// Mitsubishi GX Works2 project: ZhaoQing_HuaCheng1_Debug   PLC: Q06UDEH (continued)
    
    IF Import2Conveyor2IO.xEmpty=0 AND XF5 THEN
    	Import2LoadCylinderIO.xMDIExe:=1;
    	Import2LoadCylinderIO.iDestinationPos:=2;
    	Import2Conveyor2IO.xPutInto:=0;
    END_IF;
    IF NOT XF5 THEN
    	Import2LoadCylinderIO.xMDIExe:=1;
    	Import2LoadCylinderIO.iDestinationPos:=1;	
    END_IF;
    IF LDP(TRUE, Import2LoadCylinderIO.iCurrentPos=1) THEN
    	Import2Conveyor2IO.xPutInto:=1;
    END_IF;
   (*空框回流*)
    (*A内衬空框回流*) 
   IF  LDP(TRUE,H2200Switch1TaskID=1) THEN
   	m_xCartonADischargeLock:=1;(*A内衬空框回流下料锁，保证一次下料任务只下一个料*) 
   END_IF;
   IF LDF(TRUE,H2200BayCylinderEmptyABackIO.xUnload) OR H2200Switch1TaskID=0  THEN
   	m_xCartonADischargeLock:=0;
   END_IF;
   H2200BayCylinderEmptyABackIO.xUnload:=H2200SwitchEmptyABackConveyorIn.xEmpty
   																				 AND  H2200Switch1ConveyorIn.xEmpty
   																				 AND m_xCartonADischargeLock;
   H2200SwitchEmptyABackIO.xEntryEnable:=H2200BayCylinderEmptyABackIO.xNextRun;
   H2200SwitchEmptyABackIO.xLiftCylinderExtendInit:=H2200Switch1TaskID=1;
    H2200SwitchEmptyABackIO.xSwithEnable:=1;
    (*B内衬空框回流*) 
    IF  LDP(TRUE,H2200Switch1TaskID=2) THEN
   	m_xCartonBDischargeLock:=1;(*B内衬空框回流下料锁，保证一次下料任务只下一个料*) 
   END_IF;
   IF LDF(TRUE,H2200BayCylinderEmptyBBackIO.xUnload) OR H2200Switch1TaskID=0  THEN
   	m_xCartonBDischargeLock:=0;
   END_IF;
   H2200BayCylinderEmptyBBackIO.xUnload:=H2200SwitchEmptyBBackConveyorIn.xEmpty 
   																				 AND  H2200Switch1ConveyorIn.xEmpty
   																				 AND m_xCartonBDischargeLock;
   H2200SwitchEmptyBBackIO.xEntryEnable:=H2200BayCylinderEmptyBBackIO.xNextRun;
   H2200SwitchEmptyBBackIO.xLiftCylinderExtendInit:=1;
    H2200SwitchEmptyBBackIO.xSwithEnable:=1;    
    (*H2200Switch1 空框去注液任务*)
    IF H2200Switch1TaskID=1 OR H2200Switch1TaskID=2  THEN
    	H2200SwitchEmptyABackIO.xExitEnable:=H2200Switch1ConveyorIn.xEmpty; 
    	H2200SwitchEmptyBBackIO.xExitEnable:=H2200Switch1ConveyorIn.xEmpty;   	
    	H2200Switch1IO.xEntryEnable:=H2200SwitchEmptyABackConveyorOut.xNextRun OR H2200SwitchEmptyBBackConveyorOut.xNextRun ;
    	H2200Switch1IO.xSwithEnable:=0;
    	H2200Switch1IO.xExitEnable:=H2200RotorConveyorIO.xEmpty AND H2200RotorIO.iCurrentPos=1 AND X75;
    ELSE
    	H2200Switch1IO.xEntryEnable:=0;
    	H2200SwitchEmptyABackIO.xExitEnable:=0;
    	H2200SwitchEmptyBBackIO.xExitEnable:=0;
    	H2200Switch1IO.xExitEnable:=0;
    END_IF;
    (*H2200Switch1 满框入库任务*)
    IF H2200Switch1TaskID<>5 THEN
    	H2200Switch1IO.xLiftCylinderExtendInit:=0;
    END_IF;
    IF H2200RotorConveyorIO.xEmpty THEN
    	H2200RotorIO.xMDIExe:=1;
    	H2200RotorIO.iDestinationPos:=1;
    END_IF;
    IF H2200RotorConveyorIO.xEmpty=0 THEN
     	H2200RotorIO.xMDIExe:=1;
    	H2200RotorIO.iDestinationPos:=2;   
    END_IF;   
    IF H2200RotorIO.iCurrentPos=1 AND X75 THEN
    	H2200RotorConveyorIO.xLoad:=H2200Switch1ConveyorIn.xNextRun;
    ELSE
    	H2200RotorConveyorIO.xLoad:=0;	
    END_IF;
    IF Conveyor1IO.xEmpty THEN
    	Lifter1IO.xMDIExe:=1;
    	Lifter1IO.iDestinationPos:=2;
    END_IF;
    IF Conveyor1IO.xEmpty=0 THEN
    	Lifter1IO.xMDIExe:=1;
    	Lifter1IO.iDestinationPos:=1; 
    END_IF;
    H2200RotorConveyorIO.xUnloadCCW:=1;
    IF Lifter1IO.iCurrentPos=2 AND X8D AND H2200RotorIO.iCurrentPos=2 AND X6F THEN
    	H2200RotorConveyorIO.xUnload:=Conveyor1IO.xEmpty;
    ELSE
    	H2200RotorConveyorIO.xUnload:=0;
    END_IF;
    Conveyor1IO.xLoad:=H2200RotorConveyorIO.xNextRun; 
    IF Lifter1IO.iCurrentPos=1 AND X8C THEN
    	Conveyor1IO.xUnload:=H850Conveyor3IO.xEmpty;
    ELSE
    	Conveyor1IO.xUnload:=0;
    END_IF;  	
    H850Conveyor3IO.xLoad:=Conveyor1IO.xNextRun;
    h850conveyor3IO.xUnload:=H850Conveyor1IO.xEmpty;
    H850Conveyor1IO.xLoad:=H850Conveyor3IO.xNextRun;
    H850Conveyor1IO.xPutInto:=NOT H850Conveyor1IO.xBusy AND  SM412;
END_IF;
Y1B1:=M134 AND g_xEStop;(*空框A回流倍速链*)
Y1B0:=M135 AND g_xEStop;(*空框B回流倍速链*)
IF g_xManual THEN
    D201:=0;(*发送给化成B柜*)
    (************发送给上位机程序复位**************)
    D3100:=0;
    D3105:=0;
    D3120:=0;
    D3125:=0;
    D3016:=0;
    D3011:=0;
    D3300:=0;
    D3305:=0;
    D3310:=0;
    (*****************************************************)
	IF M163 THEN (*入库倍速链 手动*)
		 Y186:=1;(*入库倍速链*)
	ELSE
		Y186:=0;(*入库倍速链*)
	END_IF;
	IF M64 THEN (*出库倍速链 手动*)
		 Y187:=1;(*出库倍速链 *)
	ELSE
		Y187:=0;(*出库倍速链 *)
	END_IF;		
END_IF;


    (*报警*)
    M300:=NOT H3000SwitchPackageConveyorIn.xEmpty;
    M301:=H3000SwitchPackageConveyorIn.xUnloadAlarm;
    M302:=NOT H3000SwitchPackageConveyorOut.xEmpty;
    M303:=H3000SwitchPackageConveyorOut.xUnloadAlarm;   
    M304:=NOT H3000SwitchChemConveyorIn.xEmpty;
    M305:=H3000SwitchChemConveyorIn.xUnloadAlarm;   
    M306:=NOT H3000SwitchChemConveyorOut.xEmpty;
    M307:=H3000SwitchChemConveyorOut.xUnloadAlarm;  
    M308:=NOT H3000Conveyor1IO.xEmpty;
    M309:=H3000Conveyor1IO.xUnloadAlarm;       
     M310:=NOT H3000Conveyor2IO.xEmpty;
    M311:=H3000Conveyor2IO.xUnloadAlarm;    
    M312:=NOT H3000Conveyor3IO.xEmpty;
    M313:=H3000Conveyor3IO.xUnloadAlarm; 
    M314:=NOT H3000Conveyor4IO.xEmpty;
    M315:=H3000Conveyor4IO.xUnloadAlarm;  
    M317:=NOT H3000Conveyor5IO.xEmpty;
    M318:=H3000Conveyor5IO.xUnloadAlarm; 
    M319:=NOT H3000Conveyor6IO.xEmpty;
    M320:=H3000Conveyor6IO.xUnloadAlarm;     
    M321:=NOT H3000Conveyor7IO.xEmpty;
    M322:=H3000Conveyor7IO.xUnloadAlarm;  
    M323:=NOT H3000Conveyor8IO.xEmpty;
    M324:=H3000Conveyor8IO.xUnloadAlarm;  
    M325:=NOT H3000Conveyor9IO.xEmpty;
    M326:=H3000Conveyor9IO.xUnloadAlarm;  
    M327:=NOT H3000Conveyor10IO.xEmpty;
    M328:=H3000Conveyor10IO.xUnloadAlarm;
    
    M329:=NOT H3000ChemConveyor2IO.xEmpty;
    M330:=H3000ChemConveyor2IO.xUnloadAlarm;
    M331:=NOT H3000ChemConveyor3IO.xEmpty;
    M332:=H3000ChemConveyor3IO.xUnloadAlarm;
    M333:=NOT H2200Switch1ConveyorIn.xEmpty;
    M334:=H2200Switch1ConveyorIn.xUnloadAlarm;
    M335:=NOT H2200Switch1ConveyorOut.xEmpty;
    M336:=H2200Switch1ConveyorOut.xUnloadAlarm;
    M337:=NOT H2200Switch2ConveyorIn.xEmpty;
    M338:=H2200Switch2ConveyorIn.xUnloadAlarm;
    M339:=NOT H2200Switch2ConveyorOut.xEmpty;
(*    M340:=H2200Switch2ConveyorOut.xUnloadAlarm;*)
     M341:=NOT H2200Conveyor1IO.xEmpty;
    M342:=H2200Conveyor1IO.xUnloadAlarm;       
     M343:=NOT H2200Conveyor2IO.xEmpty;
    M344:=H2200Conveyor2IO.xUnloadAlarm;    
    M345:=NOT H2200Conveyor3IO.xEmpty;
    M346:=H2200Conveyor3IO.xUnloadAlarm; 
    M347:=NOT H2200Conveyor4IO.xEmpty;
    M348:=H2200Conveyor4IO.xUnloadAlarm;  
    M349:=NOT H2200Conveyor5IO.xEmpty;
    M350:=H2200Conveyor5IO.xUnloadAlarm; 
    M351:=NOT H2200Conveyor6IO.xEmpty;
    M352:=H2200Conveyor6IO.xUnloadAlarm;     
    M353:=NOT H2200Conveyor7IO.xEmpty;
    M354:=H2200Conveyor7IO.xUnloadAlarm;  
    M355:=NOT H2200Conveyor8IO.xEmpty;
    M356:=H2200Conveyor8IO.xUnloadAlarm;  
    M357:=NOT H2200Conveyor9IO.xEmpty;
    M358:=H2200Conveyor9IO.xUnloadAlarm;  
    M359:=NOT H2200Conveyor10IO.xEmpty;
    M360:=H2200Conveyor10IO.xUnloadAlarm;
    M361:=NOT H2200ImportConveyor1IO.xEmpty;
    M362:=H2200ImportConveyor1IO.xUnloadAlarm;
     M363:=NOT H2200ImportConveyor2IO.xEmpty;
    M364:=H2200ImportConveyor2IO.xUnloadAlarm;   
     M365:=NOT H2200ImportConveyor3IO.xEmpty;
    M366:=H2200ImportConveyor3IO.xUnloadAlarm;    
    M367:=NOT H850Conveyor1IO.xEmpty;
    M368:=H850Conveyor1IO.xUnloadAlarm;      
     M369:=NOT H850Conveyor3IO.xEmpty;
    M370:=H850Conveyor3IO.xUnloadAlarm;  
    M371:=NOT H850Conveyor4IO.xEmpty;
    M372:=H850Conveyor4IO.xUnloadAlarm;
    M373:=NOT H850Conveyor5IO.xEmpty;
    M374:=H850Conveyor5IO.xUnloadAlarm;
    M375:=NOT H850Conveyor6IO.xEmpty;
    M376:=H850Conveyor6IO.xUnloadAlarm;
    M377:=NOT H850Conveyor7IO.xEmpty;
    M378:=H850Conveyor7IO.xUnloadAlarm; 
    M379:=NOT H850Conveyor8IO.xEmpty;
    M380:=H850Conveyor8IO.xUnloadAlarm; 
    M381:=NOT H850RotorConveyorIO.xEmpty;
    M382:=H850RotorConveyorIO.xUnloadAlarm;     
     
    M383:=D2335=1;(*化成入库后站台读码失败*)
    M384:=D2335=3;(*化成入库后站台条码重复*)
    M385:=D2340=1;(*注液入库前站台读码失败*)
    M386:=D2340=3;(*注液入库前站台条码重复*)
    M387:=D2300=1;(*高温入库分流读码失败*)
    M388:=D2305=1;(*高温出库分流读码失败*)
    M389:=D2310=1;(*提升机2分流读码失败*)
    M390:=Lifter2IO.xLooseAlarm;(*提升机2松绳检测*)
    M391:=Conveyor2IO.xOverWidthAlarm;(*提升机2超宽报警*)
    
    M392:=Import1SwitchConveyorOut.xUnloadAlarm;
    M393:=Import2SwitchConveyorOut.xUnloadAlarm;
    M394:=NOT H1000Conveyor1IO.xEmpty;
    M395:=H1000Conveyor1IO.xUnloadAlarm;
    M396:=NOT H1000Conveyor2IO.xEmpty;
    M397:=H1000Conveyor2IO.xUnloadAlarm;
    M398:=NOT H1000Conveyor3IO.xEmpty;
    M399:=H1000Conveyor3IO.xUnloadAlarm;
    M400:=NOT H1000Conveyor4IO.xEmpty;
    M401:=H1000Conveyor4IO.xUnloadAlarm;
    M402:=NOT H1000Conveyor5IO.xEmpty;
    M403:=H1000Conveyor5IO.xUnloadAlarm;
    M404:=NOT H1000Conveyor6IO.xEmpty;
    M405:=H1000Conveyor6IO.xUnloadAlarm;
    M406:=NOT H1000Conveyor7IO.xEmpty;
    M407:=H1000Conveyor7IO.xUnloadAlarm;
    M408:=NOT H1000Conveyor8IO.xEmpty;
    M409:=H1000Conveyor8IO.xUnloadAlarm;
    M410:=NOT H1000Conveyor9IO.xEmpty;
    M411:=H1000Conveyor9IO.xUnloadAlarm;
    M412:=NOT H1000Conveyor10IO.xEmpty;
    M413:=H1000Conveyor10IO.xUnloadAlarm;
    M414:=Export1Conveyor1IO.xUnloadAlarm;
    M415:= Export2Conveyor1IO.xUnloadAlarm;
     M416:=Export1Conveyor2IO.xUnloadAlarm;
    M417:= Export2Conveyor2IO.xUnloadAlarm;   
    M418:=H850SwitchConveyorOut.xUnloadAlarm;
    g_xAlarm:=M383 
    					OR M384 
    					OR M385 
    					OR M386 
    					OR M387 
    					OR M388 
    					OR M389 
    					OR M390 
    					OR M391 
    					OR  M307 
    					OR M382 
    					OR M392 
    					OR M393 
    					OR M362
    					OR M336
    					OR M414
    					OR M415
    					OR M416
    					OR M417
    					OR M418;
  IF LDP(TRUE, g_xManual) THEN
  	m_iExportConveyorOcuppy:=0;
  END_IF;
END_PROGRAM

FUNCTION_BLOCK PriorityFB
VAR_INPUT
  xCondition1 : BOOL;  (* 条件1 *)
  xCondition2 : BOOL;  (* 条件2 *)
  xCondition3 : BOOL;  (* 条件3 *)
  xCondition4 : BOOL;  (* 条件4 *)
  xCondition5 : BOOL;  (* 条件5 *)
  xTaskComplete : BOOL;  (* 任务完成 *)
  xReset : BOOL;  (* 复位 *)
END_VAR
VAR
  xOccupy : BOOL;  (* 占用 *)
END_VAR
VAR_OUTPUT
  iPriority : INT;  (* 输出任务号 *)
END_VAR
VAR
  m_tonConditionDelay : TON;
  m_xConditionDelay : BOOL;
  m_tConditionCurrentTime : TIME;
  m_iLastTask : INT;  (* 上次执行的任务 *)
  m_tpLastTaskPulse1 : TP;
  m_xLastTaskPulse : ARRAY [1..5] OF BOOL;
  m_tLastTaskPulse : ARRAY [1..5] OF TIME := [5(T#0s)];
  m_tpLastTaskPulse2 : TP;
  m_tpLastTaskPulse3 : TP;
  m_tpLastTaskPulse4 : TP;
  m_tpLastTaskPulse5 : TP;
END_VAR
(*我在reset那里加了Occupy的复位
任务为0时，Occupy也会自动复位
*)
IF NOT xCondition1 
	AND NOT xCondition2
	AND NOT xCondition3
	AND NOT xCondition4
	AND NOT xCondition5
	AND NOT xOccupy  THEN
	iPriority:=0;
END_IF;
IF LDP(TRUE, xTaskComplete) THEN
	xOccupy:=0;
	iPriority:=0;
END_IF;
m_tonConditionDelay(IN:= (xCondition1
                                                     OR  xCondition2
                                                     OR  xCondition3
                                                     OR  xCondition4
                                                     OR xCondition5)
                                                     AND iPriority=0,
                                                     PT:= T#1s,
                                                     Q:= m_xConditionDelay ,
                                                     ET:= m_tConditionCurrentTime );
m_tpLastTaskPulse1(IN:= xCondition1  AND m_iLastTask=1 AND m_xConditionDelay  ,PT:= T#1s,Q:= m_xLastTaskPulse[1],ET:= m_tLastTaskPulse[1] );
m_tpLastTaskPulse2(IN:= xCondition2  AND m_iLastTask=2 AND m_xConditionDelay,PT:= T#1s,Q:= m_xLastTaskPulse[2],ET:= m_tLastTaskPulse[2]);
m_tpLastTaskPulse3(IN:= xCondition3  AND m_iLastTask=3 AND m_xConditionDelay,PT:= T#1s,Q:= m_xLastTaskPulse[3],ET:= m_tLastTaskPulse[3] );
m_tpLastTaskPulse4(IN:= xCondition4  AND m_iLastTask=4 AND m_xConditionDelay,PT:= T#1s,Q:= m_xLastTaskPulse[4],ET:= m_tLastTaskPulse[4] );
m_tpLastTaskPulse5(IN:= xCondition5  AND m_iLastTask=5 AND m_xConditionDelay,PT:= T#1s,Q:= m_xLastTaskPulse[5],ET:= m_tLastTaskPulse[5] );

                                                     
IF xCondition1 AND NOT xOccupy AND m_xConditionDelay AND NOT  m_xLastTaskPulse[1]  THEN
	iPriority:=1;
	xOccupy:=1;
	m_iLastTask:=1;
END_IF;
IF xCondition2 AND NOT xOccupy AND m_xConditionDelay AND NOT  m_xLastTaskPulse[2]   THEN
	iPriority:=2;
	xOccupy:=1;
	m_iLastTask:=2;
END_IF;
IF xCondition3 AND NOT xOccupy AND m_xConditionDelay AND NOT  m_xLastTaskPulse[3]   THEN
	iPriority:=3;
	xOccupy:=1;
	m_iLastTask:=3;
END_IF;
IF xCondition4 AND NOT xOccupy AND m_xConditionDelay AND NOT  m_xLastTaskPulse[4]   THEN
	iPriority:=4;
	xOccupy:=1;
	m_iLastTask:=4;
END_IF;
IF xCondition5 AND NOT xOccupy AND m_xConditionDelay AND NOT  m_xLastTaskPulse[5]   THEN
	iPriority:=5;
	xOccupy:=1;
	m_iLastTask:=5;
END_IF;

IF xReset THEN
	iPriority:=0;
	xOccupy:=0;
	m_iLastTask:=0;	
END_IF;
IF iPriority=0 THEN
	xOccupy:=0;
END_IF;
END_FUNCTION_BLOCK

FUNCTION ShuttleCarCurrentPosition
VAR_INPUT
  xPosition1 : BOOL;
  xPosition2 : BOOL;
  xPosition3 : BOOL;
END_VAR
(************************************
计算输送车当前位置的函数
**************************************)
IF xPosition1 THEN
	ShuttleCarCurrentPosition:=1;
END_IF;
IF xPosition2 THEN
	ShuttleCarCurrentPosition:=2;
END_IF;
IF xPosition3 THEN
	ShuttleCarCurrentPosition:=3;
END_IF;
END_FUNCTION

FUNCTION ShuttleCarVelocityEncoder
VAR_INPUT
  iDestinationPos : INT;  (* 目标位置 *)
  iCurrentPos : INT;  (* 当前位置 *)
  xEnable : BOOL;  (* 使能 *)
END_VAR
IF xEnable THEN
	IF ABS(iCurrentPos-iDestinationPos)<400  THEN
		ShuttleCarVelocityEncoder:=0;
	ELSE
		ShuttleCarVelocityEncoder:=1;
	END_IF;
ELSE
	ShuttleCarVelocityEncoder:=0;
END_IF;
END_FUNCTION

FUNCTION_BLOCK ShuttleCarVelocityFB
VAR_INPUT
  xEnable : BOOL;  (* 使能 *)
  xMotorCW : BOOL;  (* 电机正转 *)
  xMotorCCW : BOOL;  (* 电机反转 *)
  xPosition1Switch : BOOL;  (* 位置1开关 *)
  xDecelerationSwitch : BOOL;  (* 减速开关 *)
  xPosition2Switch : BOOL;  (* 位置2开关 *)
END_VAR
VAR
  iFloor : INT;  (* 层数 *)
END_VAR
VAR_OUTPUT
  xHighSpeed : BOOL;
END_VAR
IF xEnable THEN
	(*电机旋转，并且在位置开关上的时候触发加速*)
	IF( LDP(TRUE,xMotorCW) AND xPosition1Switch ) OR (  LDP(TRUE,xMotorCCW) AND xPosition2Switch) THEN
		xHighSpeed:=1;
		iFloor:=0;
	END_IF;
	IF LDF(TRUE,xMotorCW) OR LDF(TRUE,xMotorCCW) THEN
		xHighSpeed:=0;
    END_IF;
	IF LDP(TRUE,xDecelerationSwitch) THEN
		iFloor:=iFloor+1;
	END_IF;
	IF iFloor=2 THEN
		xHighSpeed:=0;
		iFloor:=0;
	END_IF;
ELSE
    xHighSpeed:=0;
END_IF;
END_FUNCTION_BLOCK

PROGRAM Start
IF g_xReset THEN
	SM50:=1;
ELSE
	SM50:=0;
END_IF;
CASE g_iState OF
	0: 
		g_xManual:=1;
		g_xAuto:=0;	
		g_xStackLampAmber:=1;
		g_xStackLampGreen:=0;
		g_xRemoteAuto:=0;
	1:
		g_xManual:=0;
		g_xAuto:=1;
		g_xStackLampGreen:=1;
		g_xStackLampAmber:=0;
		g_xRemoteAuto:=0;
	2:	
        g_xRemoteAuto:=1;
        g_xStackLampGreen:=1;
        g_xStackLampAmber:=0;
        g_xAuto:=0;
		g_xManual:=0;
END_CASE;
IF g_xLocalAutoStart THEN  
	g_iState:=1;
END_IF;
IF g_xAlarm AND SM412 THEN
	g_xStackLampRed:=1;
	g_xBuzzer:=1;
ELSE
	g_xStackLampRed:=0;
	g_xBuzzer:=0;	
END_IF;
IF g_xStop OR g_xEStop=0 THEN 
	g_iState:=0;
END_IF;
IF g_xRemoteAutoStart THEN
	g_iState:=2;
END_IF;
IF g_xPause AND SM412 THEN
	g_xStackLampGreen:=0;
	g_xStackLampAmber:=0;
END_IF;
END_PROGRAM

FUNCTION_BLOCK Switch
VAR_IN_OUT
  ConveyorEntryIO : ConveyorIO;
END_VAR
VAR
  ConveyorEntry : Conveyor;
END_VAR
VAR_IN_OUT
  ConveyorExitIO : ConveyorIO;
END_VAR
VAR
  m_tonLiftCylinderDelay : TON;  (* 顶升延时 *)
  m_xLiftCylinderDelay : BOOL;
  m_tLiftCylinderDelay : TIME;
  m_tonExitBarDelay : TON;  (* 退出阻挡器延时 *)
  m_tExitBarDelay : TIME;
  m_xExitBarDelay : BOOL;
END_VAR
VAR_IN_OUT
  SwitchIO : SwitchIO;
END_VAR
VAR
  iStep : INT;
  ConveyorExit : Conveyor;
  m_xInitial : BOOL;
END_VAR
(**************************************************
顶升移载模块，抽象为一条输入输线 ，一条输出输送线
一个进入阻挡器，一个放出阻挡器，和一个顶升气缸的控制
程序思路比较混乱，接口不清晰，需要整改
直接放行的时候有问题
switchEnable =0的时候   离开线体的PutInto有问题
12-17日   V1.0
***************************************************)
ConveyorEntry(ConveyorMotor:=ConveyorEntryIO);
ConveyorExit(ConveyorMotor:=ConveyorExitIO);

IF NOT m_xInitial THEN
	
	m_xInitial:=1;
END_IF;
IF g_xAuto THEN
	CASE iStep OF
		0:(*初始化*)
		ConveyorEntryIO.xLoad:=0;
		ConveyorEntryIO.xUnload:=0;
		ConveyorEntryIO.xPutInto:=0;
		ConveyorExitIO.xLoad:=0;
		ConveyorExitIo.xUnload:=0;
		ConveyorExitIO.xPutInto:=0;
		SwitchIO.xEntryBarCylinderRetract:=0;
		SwitchIO.xExitBarCylinderRetract:=0;
		IF SwitchIO.xLiftCylinderExtendInit THEN
			SwitchIO.xLiftCylinderExtend:=1;
			SwitchIO.xLiftCylinderRetract:=0;
		    IF SwitchIO.xLiftCylinderExtendDetect THEN
			    iStep:=1;
		     END_IF; 
		ELSE
			SwitchIO.xLiftCylinderExtend:=0;
			SwitchIO.xLiftCylinderRetract:=1;	
		    IF SwitchIO.xLiftCylinderRetractDetect THEN
			    iStep:=1;
		    END_IF;		
		END_IF;
		1:(*上料*)
        IF SwitchIO.xEntryEnable AND ConveyorEntryIO.xEmpty AND ConveyorExitIO.xEmpty THEN
        	SwitchIO.xEntryBarCylinderRetract:=1;
        	ConveyorEntryIO.xLoad:=1;
        END_IF;
        IF ConveyorEntryIO.xEmpty=0 THEN
        	SwitchIO.xEntryBarCylinderRetract:=0;
        	ConveyorEntryIO.xLoad:=0;
        	ConveyorExitIO.xPutInto:=1;
        END_IF;
        IF m_xLiftCylinderDelay AND  SwitchIO.xSwithEnable THEN
        	 iStep:=2;
        END_IF;
        IF SwitchIO.xSwithEnable=0 AND m_xLiftCylinderDelay  THEN
        	 iStep:=3;
        END_IF;
		2:(*顶升*)
			SwitchIO.xExitBarCylinderRetract:=0;
		    IF SwitchIO.xLiftCylinderExtendInit THEN
			    SwitchIO.xLiftCylinderExtend:=0;
			    SwitchIO.xLiftCylinderRetract:=1;
		    ELSE
			    SwitchIO.xLiftCylinderExtend:=1;
			    SwitchIO.xLiftCylinderRetract:=0;			
		   END_IF;

		  IF SwitchIO.xLiftCylinderExtendInit THEN
		  	IF SwitchIO.xLiftCylinderRetractDetect THEN
		  		iStep:=4;
		  	END_IF;
		  	ELSE
		  	IF SwitchIO.xLiftCylinderExtendDetect THEN
		      iStep:=4; 
		  	END_IF;
		  END_IF;
		  3:(*放行*)	
		  	SwitchIO.xExitBarCylinderRetract:=1;
		  	ConveyorExitIO.xPutInto:=0;
		  	iStep:=4;
		  4:(*下料*)
		  (*通过出料传输线下料*)
		  IF SwitchIO.xExitEnable  AND m_xExitBarDelay AND NOT SwitchIO.xExitBarCylinderRetract  THEN		  
		  	ConveyorExitIO.xUnload:=1;
		  ELSE
		  	ConveyorExitIO.xUnload:=0;
		  END_IF;	
		   (*通过进料传输线下料*)
		  IF SwitchIO.xExitEnable  AND m_xExitBarDelay  AND SwitchIO.xExitBarCylinderRetract THEN		  
		  	ConveyorEntryIO.xUnload:=1;
		  ELSE
		  	ConveyorEntryIO.xUnload:=0;
		  END_IF;			    	
		  IF ConveyorExitIO.xEmpty OR ConveyorEntryIO.xEmpty  THEN
		  	ConveyorExitIO.xPutInto:=1;
		  	ConveyorEntryIO.xPutInto:=1;
			iStep:=0; 
		  END_IF;
	END_CASE;
        m_tonLiftCylinderDelay(IN:=NOT ConveyorEntryIO.xEmpty AND iStep=1 ,PT:= T#1S ,Q:= m_xLiftCylinderDelay ,ET:=m_tLiftCylinderDelay );
 		m_tonExitBarDelay(IN:=iStep=4 ,PT:= T#1s ,Q:= m_xExitBarDelay ,ET:= m_tExitBarDelay);
END_IF;
(*复位程序*)
IF (g_xResetSingle AND  (g_iDeviceIDSelect=ConveyorEntryIO.iDeviceID OR g_iDeviceIDSelect=ConveyorExitIO.iDeviceID))
	OR LDP(TRUE,SwitchIO.xLiftCylinderExtendInit) 
	OR LDF(TRUE,SwitchIO.xLiftCylinderExtendInit) 
	 THEN
	ConveyorEntryIO.xPutInto:=1;
	ConveyorExitIO.xPutInto:=1;
	iStep:=0;
END_IF;
IF g_xManual  THEN
	iStep:=0;
	ConveyorEntryIO.xLoad:=0;
    ConveyorEntryIO.xUnload:=0;
	ConveyorEntryIO.xPutInto:=0;
	ConveyorExitIO.xLoad:=0;
	ConveyorExitIo.xUnload:=0;
	ConveyorExitIO.xPutInto:=0;
	SwitchIO.xEntryBarCylinderRetract:=0;
	SwitchIO.xExitBarCylinderRetract:=0;
	IF SwitchIO.xEntryBarCylinderRetractButton THEN
		SwitchIO.xEntryBarCylinderRetract:=1;
	ELSE
		SwitchIO.xEntryBarCylinderRetract:=0;
	END_IF;
		IF SwitchIO.xExitBarCylinderRetractButton THEN
		SwitchIO.xExitBarCylinderRetract:=1;
	ELSE
		SwitchIO.xExitBarCylinderRetract:=0;
		END_IF;
		IF SwitchIO.xLiftCylinderExtendButton AND NOT SwitchIO.xLiftCylinderRetractButton THEN
			SwitchIO.xLiftCylinderExtend:=1;
			SwitchIO.xLiftCylinderRetract:=0;
		END_IF;
		IF NOT SwitchIO.xLiftCylinderExtendButton AND  SwitchIO.xLiftCylinderRetractButton THEN
			SwitchIO.xLiftCylinderExtend:=0;
			SwitchIO.xLiftCylinderRetract:=1;
		END_IF;		
	END_IF;
END_FUNCTION_BLOCK

PROGRAM UDP
VAR
  m_ton1ReceiveHeartbeat : TON;
  m_t1RecHeartbeatCurrentTime : TIME;
  m_tonAutoClose : TON;
  m_xAutoClose : BOOL;
  m_tAutoCloseCurrentTime : TIME;
  m_tonReconnect : TON;
  m_xReconnect : BOOL;
  m_tReconnectCurrentTime : TIME;
  m_ton5ReceiveHeartbeat : TON;
  m_t5RecHeartbeatCurrentTime : TIME;
END_VAR
(*与化成柜2通讯*)
D200:=2;
m_tonReconnect(IN:= NOT SD1282.0 AND NOT SD1284.0,PT:=T#5s  ,Q:=m_xReconnect ,ET:=m_tReconnectCurrentTime);
SP_SOCOPEN(m_xReconnect  AND SD1288.A , "U0", K1 , D110 , M100);
SP_SOCSND( SM412 AND SD1282.0 , "U0" , K1 , D100, D200, M102 );
SP_SOCRCV( SD1282.0 AND SD1286.0 AND NOT M104 , "U0" , K1, D300 , D400 ,M104 );
m_tonAutoClose(IN:= SD1284.0 AND NOT SD1282.0 ,PT:=T#5s,Q:=m_xAutoClose ,ET:= m_tAutoCloseCurrentTime );
SP_SOCCLOSE( LDF(TRUE,SD1282.0) OR m_xAutoClose  , "U0" , K1, D120, M106 );
D201.F:=SM413;
m_ton1ReceiveHeartbeat(IN:=NOT LDP(TRUE, D401.F) ,PT:= t#5S ,Q:= g_xChem2ComFailed ,ET:= m_t1RecHeartbeatCurrentTime);
IF g_xChem2ComFailed THEN
	M104:=SM413;(*通讯失败有可能是接收模块没动作，重启接收模块*)
	D400:=0;
	D401:=0;
END_IF;
(*编码器处理程序*)
IF XA OR X0B   THEN
	D140:=2;
	D143:=6;
END_IF;
	G_INPUT( X0A OR X0B AND NOT M110, 0 , D140 , D160 , M110 );(*串口数据读取指令*)
(*IF M110 THEN
	D170:=0;
	D172:=4;
END_IF;*)
(*使用可变长度报文，通过接收结束代码的接收方法，默认的是CR+LF
编码器只发CR，需要在智能模块中设置成CR为结束符，这样不需要ZP_CSET指令清除串口缓存区*)
(*ZP_CSET( M110  , "U0", 2 , D170, D180,M112 );(*串口数据缓存区清除指令*)
IF D160=11069 THEN  (*接收到数据开始执行ASCII码转换成10进制，D160为=+ ，串口传输的字头 转换为10进制是11069，不判断这个报4100错误*)
    DABIN( TRUE , D163, D190 );
END_IF;

(*注液RGV，TCP通讯*)
D240:=k8;
SP_SOCCINF( LDP(TRUE,SD1282.4) , "U0" , K5 , D500 ,D520);
SP_SOCSND( SM412 AND SD1282.4 , "U0" , K5 , D510, D240, M114);
SP_SOCRCV( NOT M116 AND SD1282.4 , "U0" , K5, D320 , D440 ,M116);
D243.F:=SM413;
m_ton5ReceiveHeartbeat(IN:=NOT LDP(TRUE, D443.F) ,PT:= t#5S ,Q:= g_xFillingRGVComFailed ,ET:= m_t5RecHeartbeatCurrentTime);
END_PROGRAM

FUNCTION_BLOCK Conveyor
VAR
  tRundelay : TIME;  (* 离开延时 *)
END_VAR
VAR_IN_OUT
  ConveyorMotor : ConveyorIO;  (* 输送线输入输出 *)
END_VAR
VAR
  iStep : INT;  (* 上料步骤 *)
  m_tUnloadTimer : TIME;  (* 下料计时器 *)
  m_tonLeaveDelay : TON;  (* 离开延时定时器 *)
  m_xLeaveDelayOut : BOOL;  (* 离开延时 *)
  m_tLeaveCurrentTime : TIME;
END_VAR
VAR CONSTANT
  LOAD_UNLOAD_TIME : TIME := T#30s;  (* 延时报警常量 *)
END_VAR
VAR
  m_tonUnloadAlam : TON;  (* 下料报警定时器 *)
  m_tonLoadDelay : TON;  (* 离开延时定时器 *)
  m_xLoadDelayOut : BOOL;  (* 离开延时 *)
  m_tLoadCurrentTime : TIME;
  m_xInitial : BOOL;  (* 初始化 *)
  m_tLoadTimer : TIME;  (* 上料延时当前时间 *)
END_VAR
(*////////////////////////////////////////////////////////////////////////////////////////////////////////////
//传输线控制FB块，可控制单方向线体，双向旋转线体，支持双向上下料            
//线体初始化后为空的情况下输入xLoad信号即可进行上料动作，使用xLoadCCW信号可反方向上料
//增加了产品信息和产品种类的储存，当传输线为空和上料进行标志位为零的情况下清除产品信息和产品种类
//使用方式是在置位xLoad信号后，把产品信息和产品种类传入，等下料后自动清零
//线体不为空的情况下使用xUnload信号可进行下料动作，物料有无传感器的下降沿后出发计时器，延时断开传输线旋转
//单方向传输线体把xLoadCCW、xUnloadCCW设置为零，双向线体上料方向和下料反向的,方向固定的 把xUnloadCCW设置为1
//双方向线体双向都能上下料的要根据上料的方向来设置xLoadCCW,xUnloadCCW
//增加工作中信号xBusy当电机正转 显示为工作中
//增加上下料超时报警，xLoadAlarm，xUnloadAlarm，设定时间在LOAD_UNLOAD_TIME常量上，现在设置的为30秒
//增加xPutInto信号，用于直接投入的物料，检测开关感应到后，直接进入下料流程，上升沿有效
//离开延时改为变量 iLeaveDelay 默认为0 离开检测开关离输送线尾端比较远的线体需要根据情况设定100ms为单位
增加初始化标志位，增加进入延时时间，初始化为进入延时时间为0 ，离开延时时间为2S，通过外围接口可以更改
//修改信息  修改后请增加版本
//YAO      V1.0
///////////////////////////////////////////////////////////////////////////////////////////////////////////
********************************************************)
IF NOT m_xInitial THEN
	ConveyorMotor.tLoadDelay:=T#100ms;
	ConveyorMotor.xNegLimit:=1;
	ConveyorMotor.xPosLimit:=1;
	ConveyorMotor.xSizeDeficientDetect:=0;
END_IF;
m_xInitial:=1;
IF g_xAuto THEN
CASE iStep OF
	0:
	ConveyorMotor.xMotorCW:=0;
	ConveyorMotor.xMotorCCW:=0;
	ConveyorMotor.xNextRun:=0;
IF g_xEStop AND NOT ConveyorMotor.xLimitAlarrm AND NOT ConveyorMotor.xOverWidthAlarm  THEN
	IF  ConveyorMotor.xCWPresent OR ConveyorMotor.xCCWPresent  THEN
		iStep:=3;
		ConveyorMotor.xEmpty:=0;
		ELSE
		iStep:=1;
		ConveyorMotor.xEmpty:=1;
	END_IF;
END_IF;		
	1: 
	IF ConveyorMotor.xLoad    
		AND ConveyorMotor.xMotorCW=0   
		AND ConveyorMotor.xMotorCCW=0   
		AND ConveyorMotor.xEmpty THEN	
		iStep:=2;
	END_IF;
	2: 
	IF ConveyorMotor.xloadCCW THEN
		ConveyorMotor.xMotorCCW:=1; 
		ConveyorMotor.xMotorCW:=0;
	ELSE
	    ConveyorMotor.xMotorCW:=1;  
		ConveyorMotor.xMotorCCW:=0;
	END_IF;
		m_tonLoadDelay(IN:= (ConveyorMotor.xCWPresent AND NOT ConveyorMotor.xloadCCW) 
		                                        OR (ConveyorMotor.xCCWPresent AND ConveyorMotor.xloadCCW) ,
		                               PT:= ConveyorMotor.tLoadDelay ,
		                               Q:= m_xLoadDelayOut ,
		                               ET:= m_tLoadTimer );
	    IF (m_xLoadDelayOut AND NOT ConveyorMotor.xSizeDeficientDetect)   (*无尺寸检测时  只检测一个开关*)
	    	OR (m_xLoadDelayOut AND ConveyorMotor.xSizeDeficientDetect(*有尺寸检测时  要检测两个开关*)
	    	                                          AND ConveyorMotor.xCCWPresent 
	    	                                          AND ConveyorMotor.xCWPresent)      THEN 	 
		    iStep:=3;
			    ELSIF (m_xLoadDelayOut 
		                       AND ConveyorMotor.xSizeDeficientDetect(*尺寸不足报警*)
	    	                  AND (NOT ConveyorMotor.xCCWPresent OR NOT ConveyorMotor.xCWPresent))  
	    THEN
	    	    ConveyorMotor.xOverWidthAlarm:=1;
	    	   iStep:=0;               
	    END_IF;
	    
	3:
	ConveyorMotor.xMotorCW:=0;
	ConveyorMotor.xMotorCCW:=0;
	ConveyorMotor.xEmpty:=0;
	IF ConveyorMotor.xUnload AND NOT ConveyorMotor.xOverWidthAlarm THEN 
		iStep:=4;
	END_IF;
	4:	
	IF ConveyorMotor.xUnloadCCW THEN   
		ConveyorMotor.xMotorCCW:=1;  
		ConveyorMotor.xMotorCW:=0;
		ELSE
	    ConveyorMotor.xMotorCW:=1;  
		ConveyorMotor.xMotorCCW:=0;
	END_IF;
	ConveyorMotor.xNextRun:=1; 
	IF NOT ConveyorMotor.xUnload THEN 
		istep:=0;
	END_IF;
END_CASE;
IF LDP(TRUE,ConveyorMotor.xPutInto) THEN
	iStep:=0;
END_IF;
END_IF;
IF g_xManual THEN
	iStep:=0;

	IF ConveyorMotor.xForward 
		AND ConveyorMotor.xBackward=0 
		AND ConveyorMotor.xMotorCCW=0
		AND g_xEStop THEN
		ConveyorMotor.xMotorCW:=1;
		ConveyorMotor.xMotorCCW:=0;
		ELSE
		ConveyorMotor.xMotorCW:=0;
	END_IF;

	IF ConveyorMotor.xBackward 
		AND ConveyorMotor.xForward=0 
		AND ConveyorMotor.xMotorCW=0
		AND g_xEStop  THEN
		ConveyorMotor.xMotorCCW:=1;
		conveyormotor.xMotorCW:=0;
		ELSE
		ConveyorMotor.xMotorCCW:=0;
	END_IF;
END_IF;
IF ConveyorMotor.xMotorCCW        
	OR ConveyorMotor.xMotorCW THEN  
	ConveyorMotor.xBusy:=1;
	ELSE
	ConveyorMotor.xBusy:=0;
END_IF;
m_tonUnloadAlam(IN:= iStep=4,PT:= LOAD_UNLOAD_TIME,Q:= ConveyorMotor.xUnloadAlarm,ET:= m_tUnloadTimer );
(*//复位*)
IF (*g_xReset OR*)
	 (g_xResetSingle AND ConveyorMotor.iDeviceID=g_iDeviceIDSelect)THEN (*AND ConveyorMotor.iDeviceID=g_iDeviceIDSelect  THEN*)  (* //非正常情况下切断xNextRun不会复位，通过这个标志位会出发报警*)(*增加单体复位*)
	iStep:=0;
	ConveyorMotor.xNextRun:=0; 
	ConveyorMotor.xLimitAlarrm:=0;
	ConveyorMotor.xOverWidthAlarm:=0;
END_IF;
IF iStep=3 AND (NOT ConveyorMotor.xNegLimit OR NOT ConveyorMotor.xPosLimit) THEN
	ConveyorMotor.xOverWidthAlarm:=1;
END_IF;
IF ( ((ConveyorMotor.xloadCCW AND NOT ConveyorMotor.xNegLimit)            (*反转上料，碰到负限位*)
	OR  ( NOT ConveyorMotor.xloadCCW AND NOT ConveyorMotor.xPosLimit)) (*正转上料，碰到正限位*)
    AND iStep=2) (*上料过程*)
    OR
   ( iStep=4 (*下料过程*)
	AND( (ConveyorMotor.xUnloadCCW AND NOT ConveyorMotor.xPosLimit)  
	OR (NOT ConveyorMotor.xUnloadCCW AND NOT ConveyorMotor.xNegLimit)))    
    THEN
    ConveyorMotor.xLimitAlarrm:=1;
    iStep:=0;
END_IF;
END_FUNCTION_BLOCK

FUNCTION_BLOCK ShuttleCar
VAR_IN_OUT
  ShuttleCarInOut : ShuttleCarIO;
END_VAR
VAR
  m_tonBrakeDelay : TON;  (* 延时 *)
  m_tBrakeDelayCurrentTime : TIME;
  m_tonArriveDelay : TON;  (* 到达延时计时器 *)
  m_xInit : BOOL;  (* 初始化标志位 *)
  m_tonPauseDelay : TON;  (* 暂停减速 *)
  m_tPauseDelayCurrentTime : TIME;  (* 暂停延时当前时间 *)
  m_xArriveDelay : BOOL;  (* 到达延时 *)
  m_tArriveDelayCurrentTime : TIME;  (* 到达延时当前时间 *)
  m_tonOvertimeAlarm : TON;  (* 超时报警定时器 *)
  m_tOvertimeCurrentTime : TIME;  (* 超时报警当前时间 *)
END_VAR
(*******************************************************************
输送小车程序，可用于使用认址片控制位置的输送车程序，可用于控制提升机，
使用了限位捕捉程序防止小车惯性过大冲过限位后继续行走，捕捉程序采用反
转复位，这样设计有弊端可能反转复位后车的位置并没有回到限位以内,当两个
限位同时碰到的时候，会使运料小车进入死锁状态，通过xPassLimit来解开死锁，
可以在触摸屏中使用一个带权限的按钮来进行控制，配合ShuttleCarCurrentPos
函数来计算位置信息
增加自动开始后将当前位置置为零的信号防止设备停在两个位置开关的中间
修改信息  修改后请增加版本
2018-1-22增加到位延时：到位延时时间可以设置，适应双向到位的位置开关，通过调整延时时间让穿梭车停在到位开关的中间
增加气缸控制信号
增加抱闸延时
增加超时报警
YAO      V1.0
2018-1-22 YAO V1.1
********************************************************************)
IF NOT m_xInit THEN
	ShuttleCarInOut.tArriveDelay:=T#0s;   (*到位延时初始化为0*)
	ShuttleCarInOut.tBrakeDelay:=T#100ms;(*抱闸延时初始化为100ms*)
	ShuttleCarInOut.tSetOverTime:=T#60s;(*超时报警初始化为1分钟*)
	m_xInit:=1;
END_IF;
(*如果是气缸的话屏蔽限位和Ready信号*)
IF ShuttleCarInOut.xCylinder THEN
	ShuttleCarInOut.xPosLimit:=1;
	ShuttleCarInOut.xNegLimit:=1;
	ShuttleCarInOut.xReady:=1;
END_IF;
(*限位捕捉，防止冲过限位开关，反转后复位*)
ShuttleCarInOut.xPosLimitCatch:=LDF(TRUE,ShuttleCarInOut.xPosLimit) OR ShuttleCarInOut.xPosLimitCatch;
IF ShuttleCarInOut.xCCW THEN  
	ShuttleCarInOut.xPosLimitCatch:=0;
END_IF;

ShuttleCarInOut.xNegLimitCatch:=LDF(TRUE,ShuttleCarInOut.xNegLimit) OR ShuttleCarInOut.xNegLimitCatch;
(*松绳报警*)
IF LDP(TRUE,ShuttleCarInOut.xLooseDetect) THEN	
	ShuttleCarInOut.xLooseAlarm:=1;
END_IF;
(*提升复位报警*)
IF ShuttleCarInOut.xCW AND NOT  ShuttleCarInOut.xLooseDetect THEN   
	ShuttleCarInOut.xLooseAlarm:=0; 
END_IF;

IF ShuttleCarInOut.xCW THEN   
	ShuttleCarInOut.xNegLimitCatch:=0; 
END_IF;

IF ShuttleCarInOut.xPassLimit OR
	g_xReset OR   (*增加复位按钮*)
	(ShuttleCarInOut.xNegLimitCatch 
	AND ShuttleCarInOut.xPosLimitCatch)  THEN  
	ShuttleCarInOut.xNegLimitCatch:=0; 
	ShuttleCarInOut.xPosLimitCatch:=0;
	ShuttleCarInOut.xLooseAlarm:=0;
END_IF;
IF ShuttleCarInOut.xReady AND g_xEStop THEN
(*手动*)
    IF g_xManual THEN  
	    IF ShuttleCarInOut.xForward 
			AND ShuttleCarInOut.xBackward=0 
			AND ShuttleCarInOut.xCCW=0 
			AND ShuttleCarInOut.xPosLimitCatch=0  THEN
		    ShuttleCarInOut.xCW:=1;
		    ELSE
		    ShuttleCarInOut.xCW:=0;
	    END_IF;
	    IF ShuttleCarInOut.xBackward 
			AND ShuttleCarInOut.xForward=0 
			AND ShuttleCarInOut.xCW=0 
			AND ShuttleCarInOut.xNegLimitCatch=0 
			AND ShuttleCarInOut.xLooseAlarm=0
			AND G_xEStop THEN  
		    ShuttleCarInOut.xCCW:=1;
		    ELSE
		    ShuttleCarInOut.xCCW:=0;
	    END_IF;
    END_IF;
    (**********)
(*自动*)
  IF g_xAuto  THEN  
  	(*点动*)
 		IF LDP(TRUE,ShuttleCarInOut.xForward) THEN
 			ShuttleCarInOut.xMDIExe:=1;
			ShuttleCarInOut.iDestinationPos:=ShuttleCarInOut.iCurrentPos+1;
		END_IF;
		IF LDP(TRUE,ShuttleCarInOut.xBackward) THEN
			ShuttleCarInOut.xMDIExe:=1;
			ShuttleCarInOut.iDestinationPos:=ShuttleCarInOut.iCurrentPos-1;
		END_IF;	 
	(*>>>>>>>>>>>>>>>>>>>>>>>>>>>>>>>>>>>>>*)	
	  IF ShuttleCarInOut.xMDIExe AND ShuttleCarInOut.iDestinationPos<>0 THEN	
	    IF ShuttleCarInOut.iCurrentPos<ShuttleCarInOut.iDestinationPos AND ShuttleCarInOut.xPosLimitCatch=0 THEN   (*正转*)
			ShuttleCarInOut.xCW:=1;
			ShuttleCarInOut.xCCW:=0;
			ShuttleCarInOut.xMDIDone:=0;
		END_IF;

		IF ShuttleCarInOut.iCurrentPos>ShuttleCarInOut.iDestinationPos AND ShuttleCarInOut.xNegLimitCatch=0 AND ShuttleCarInOut.xLooseAlarm=0 THEN   (*反转*)
			ShuttleCarInOut.xCCW:=1;
			ShuttleCarInOut.xCW:=0;
			ShuttleCarInOut.xMDIDone:=0;
		END_IF;
	m_tonArriveDelay(IN:= ShuttleCarInOut.iCurrentPos=ShuttleCarInOut.iDestinationPos ,
	                                    PT:= ShuttleCarInOut.tArriveDelay ,
	                                    Q:= m_xArriveDelay ,
	                                    ET:= m_tArriveDelayCurrentTime);
	     (*到位延时时间可以设置，适应双向到位的位置开关，通过调整延时时间让穿梭车停在到位开关的中间*)
		IF m_xArriveDelay AND NOT ShuttleCarInOut.xCylinder THEN
			ShuttleCarInOut.xCW:=0;
			ShuttleCarInOut.xCCW:=0;
			ShuttleCarInOut.xMDIDone:=1;
			ELSE
			ShuttleCarInOut.xMDIDone:=0;
		END_IF;

		IF ShuttleCarInOut.xPosLimitCatch THEN
			ShuttleCarInOut.xCW:=0;
			ShuttleCarInOut.xMDIDone:=0;
		END_IF;

		IF ShuttleCarInOut.xNegLimitCatch THEN
			ShuttleCarInOut.xCCW:=0;
			ShuttleCarInOut.xMDIDone:=0;
		END_IF;
		ELSE
		ShuttleCarInOut.xCW:=0;
		ShuttleCarInOut.xCCW:=0;
		ShuttleCarInOut.xMDIDone:=0;
	  END_IF;
	END_IF;
	ELSE  (*无就绪信号   或急停的情况下*)
		ShuttleCarInOut.xCW:=0;
		ShuttleCarInOut.xCCW:=0;	
END_IF;
    (*抱闸延时*)
m_tonBrakeDelay(IN:= ShuttleCarInOut.xCW OR ShuttleCarInOut.xCCW,
                                    PT:= ShuttleCarInOut.tBrakeDelay,
                                    Q:=ShuttleCarInOut.xBrake ,
                                    ET:= m_tBrakeDelayCurrentTime);

(*自动上电后把当前位置清零，防止穿梭车不在开关位置*)
IF LDP(TRUE,g_xAuto) THEN
	ShuttleCarInOut.iCurrentPos:=0;
END_IF;
IF ShuttleCarInOut.xCW OR ShuttleCarInOut.xCCW THEN
	ShuttleCarInOut.xBusy:=1;
	ELSE
	ShuttleCarInout.xBusy:=0;
END_IF;

(*暂停，带延时减速斜坡，ShuttleCarInOut.xPauseRamp为减速斜坡输出位*)
m_tonPauseDelay(IN:=g_xPause,PT:= T#2s ,Q:=ShuttleCarInOut.xPauseRamp,ET:= m_tPauseDelayCurrentTime );
IF ShuttleCarInOut.xPauseRamp THEN
	ShuttleCarInOut.xCW:=0;
	ShuttleCarInOut.xCCW:=0;
	ShuttleCarInOut.xBrake:=0;
END_IF;
(*超时报警*)
m_tonOvertimeAlarm(IN:= ShuttleCarInOut.xMDIExe AND (ShuttleCarInOut.iCurrentPos<>ShuttleCarInOut.iDestinationPos) ,
                                           PT:= ShuttleCarInOut.tSetOverTime,
                                           Q:= ShuttleCarInOut.xOvertimeAlarm ,
                                           ET:= m_tOvertimeCurrentTime );
END_FUNCTION_BLOCK

FUNCTION_BLOCK BarCylinder
VAR_IN_OUT
  BarCylinderIO : BarCylinderIO;
END_VAR
VAR
  m_xInitial : BOOL;  (* 初始化 *)
  m_tonLoadDelay : TON;  (* 上料延时 *)
  m_xLoadDelay : BOOL;  (* 上料延时标志位 *)
  m_tLoadDelayCurrentTime : TIME;  (* 上料延时当前时间 *)
END_VAR
  (***********************************************************************
阻挡器模块，
由一个行程开关，一个阻挡器，一个倍速链输送电机组成
具有手动与自动模式
xEmpty显示当前为空料的状态
xUnload为卸料信号，连接下一设备的xEmpty信号
增加分料气缸xBarCylinderSecondary
增加复位功能，Unload NextRun  Empty 能形成死锁，如果Unload 信号一直给，会造成无法复位
*************************************************************************)

